      ReacTi : G7_TransitionPlus_V6;   // Transition structure
      ReacD : G7_TransitionPlus_V6;   // Transition structure
      Confirm : G7_TransitionPlus_V6;   // Transition structure
      UserBtch : G7_TransitionPlus_V6;   // Transition structure
      "StT-103" : G7_TransitionPlus_V6;   // Transition structure
      Route_Ok : G7_TransitionPlus_V6;   // Transition structure
      MixDone : G7_TransitionPlus_V6;   // Transition structure
      TimeOut : G7_TransitionPlus_V6;   // Transition structure
      EmptyLv : G7_TransitionPlus_V6;   // Transition structure
      LR : G7_TransitionPlus_V6;   // Transition structure
      LFUW : G7_TransitionPlus_V6;   // Transition structure
      mtL : G7_TransitionPlus_V6;   // Transition structure
      DneTransf : G7_TransitionPlus_V6;   // Transition structure
      TWash : G7_TransitionPlus_V6;   // Transition structure
      STW : G7_TransitionPlus_V6;   // Transition structure
      OpRout : G7_TransitionPlus_V6;   // Transition structure
      TW_RW : G7_TransitionPlus_V6;   // Transition structure
      TW_Vfd : G7_TransitionPlus_V6;   // Transition structure
      Trans87 : G7_TransitionPlus_V6;   // Transition structure
      TW_Wng : G7_TransitionPlus_V6;   // Transition structure
      TW_VfdOf : G7_TransitionPlus_V6;   // Transition structure
      Trans90 : G7_TransitionPlus_V6;   // Transition structure
      DneTnkW : G7_TransitionPlus_V6;   // Transition structure
      TE_SWW : G7_TransitionPlus_V6;   // Transition structure
      TuW : G7_TransitionPlus_V6;   // Transition structure
      STuW : G7_TransitionPlus_V6;   // Transition structure
      Trans103 : G7_TransitionPlus_V6;   // Transition structure
      TuWRW : G7_TransitionPlus_V6;   // Transition structure
      TuWGW : G7_TransitionPlus_V6;   // Transition structure
      TuW_SRW : G7_TransitionPlus_V6;   // Transition structure
      TuW_R : G7_TransitionPlus_V6;   // Transition structure
      Trans108 : G7_TransitionPlus_V6;   // Transition structure
      Trans109 : G7_TransitionPlus_V6;   // Transition structure
      PmpsOn : G7_TransitionPlus_V6;   // Transition structure
      ReEmpty : G7_TransitionPlus_V6;   // Transition structure
      PmpsOff : G7_TransitionPlus_V6;   // Transition structure
      OutleClsd : G7_TransitionPlus_V6;   // Transition structure
      DneTubW : G7_TransitionPlus_V6;   // Transition structure
      Init : G7_TransitionPlus_V6;   // Transition structure
      SAut : G7_TransitionPlus_V6;   // Transition structure
      SIn : G7_TransitionPlus_V6;   // Transition structure
      Initd : G7_TransitionPlus_V6;   // Transition structure
      WaterDn : G7_TransitionPlus_V6;   // Transition structure
      Ab : G7_TransitionPlus_V6;   // Transition structure
      AbortOn : G7_TransitionPlus_V6;   // Transition structure
      DneAbort : G7_TransitionPlus_V6;   // Transition structure
      Idle : G7_StepPlus_V6;   // Step structure
      Ready : G7_StepPlus_V6;   // Step structure
      SelectSeq : G7_StepPlus_V6;   // Step structure
      Started : G7_StepPlus_V6;   // Step structure
      StartTanks : G7_StepPlus_V6;   // Step structure
      FillingUpWater : G7_StepPlus_V6;   // Step structure
      StopReqWaterP : G7_StepPlus_V6;   // Step structure
      ReleaseWTank : G7_StepPlus_V6;   // Step structure
      "Pre-Mix" : G7_StepPlus_V6;   // Step structure
      OpenRoutes : G7_StepPlus_V6;   // Step structure
      X : G7_StepPlus_V6;   // Step structure
      FillDone_T101 : G7_StepPlus_V6;   // Step structure
      Close_T101 : G7_StepPlus_V6;   // Step structure
      "T-101_Done" : G7_StepPlus_V6;   // Step structure
      Y : G7_StepPlus_V6;   // Step structure
      pH_Ctrl1 : G7_StepPlus_V6;   // Step structure
      pH_Ctrl2 : G7_StepPlus_V6;   // Step structure
      FillDone_T102 : G7_StepPlus_V6;   // Step structure
      Close_T102 : G7_StepPlus_V6;   // Step structure
      "T-102_Done" : G7_StepPlus_V6;   // Step structure
      ReactingTime : G7_StepPlus_V6;   // Step structure
      ReactingDone : G7_StepPlus_V6;   // Step structure
      "USER Waiting" : G7_StepPlus_V6;   // Step structure
      "EDIT BatchP" : G7_StepPlus_V6;   // Step structure
      "Start T-103" : G7_StepPlus_V6;   // Step structure
      "R-201-->T-103" : G7_StepPlus_V6;   // Step structure
      MixToClean : G7_StepPlus_V6;   // Step structure
      LastFlushOut : G7_StepPlus_V6;   // Step structure
      Transfering : G7_StepPlus_V6;   // Step structure
      LastFIllUp : G7_StepPlus_V6;   // Step structure
      FirstFlushOut : G7_StepPlus_V6;   // Step structure
      LastFillUpW : G7_StepPlus_V6;   // Step structure
      LastTransfer : G7_StepPlus_V6;   // Step structure
      Done_Transfer : G7_StepPlus_V6;   // Step structure
      Idle_TWash : G7_StepPlus_V6;   // Step structure
      Start_TWash : G7_StepPlus_V6;   // Step structure
      OpenRoute : G7_StepPlus_V6;   // Step structure
      ReqWaterWash : G7_StepPlus_V6;   // Step structure
      "2011 VFD ON & PID AUTO/Wait for 80%_R-201" : G7_StepPlus_V6;   // Step structure
      StopWaterWash : G7_StepPlus_V6;   // Step structure
      "XV-1043_CC_02_R-201" : G7_StepPlus_V6;   // Step structure
      Washing : G7_StepPlus_V6;   // Step structure
      "2011VFD OFF & PID MAN_R-201" : G7_StepPlus_V6;   // Step structure
      USER_MAN_DRAIN : G7_StepPlus_V6;   // Step structure
      Done_TWash : G7_StepPlus_V6;   // Step structure
      Idle_TubWash : G7_StepPlus_V6;   // Step structure
      Start_TubWash : G7_StepPlus_V6;   // Step structure
      "XV-1043_CO_03_R-201" : G7_StepPlus_V6;   // Step structure
      ReqWaterTuW : G7_StepPlus_V6;   // Step structure
      GettingWater : G7_StepPlus_V6;   // Step structure
      StopRqWaterTuW : G7_StepPlus_V6;   // Step structure
      "ReleaseT-104" : G7_StepPlus_V6;   // Step structure
      "XV-1043_CC_03_R-529" : G7_StepPlus_V6;   // Step structure
      "XV-2013_CO_XV-1043_Cc_R-201" : G7_StepPlus_V6;   // Step structure
      "P-201A/B_ON_R-201" : G7_StepPlus_V6;   // Step structure
      Emptying : G7_StepPlus_V6;   // Step structure
      "P-201A/B_OFF_R-201" : G7_StepPlus_V6;   // Step structure
      Close_Outlet : G7_StepPlus_V6;   // Step structure
      Done_TubWash : G7_StepPlus_V6;   // Step structure
      Initialize : G7_StepPlus_V6;   // Step structure
      SetAuto : G7_StepPlus_V6;   // Step structure
      SetInitial : G7_StepPlus_V6;   // Step structure
      Initialized : G7_StepPlus_V6;   // Step structure
      AbortStarting : G7_StepPlus_V6;   // Step structure
      Aborting : G7_StepPlus_V6;   // Step structure
      Abort_Done : G7_StepPlus_V6;   // Step structure
      SINI : Array[0..9] of USInt;
      LSTT : Array[0..68] of USInt;
      ATAJ : Array[0..68] of USInt;
      ATAB : Array[0..68] of USInt;
      PSTT : Array[0..68] of USInt;
      NSTT : Array[0..68] of USInt;
      ASSJ : Array[0..65] of USInt;
      ASSB : Array[0..65] of USInt;
      PTTS : Array[0..65] of USInt;
      NTTS : Array[0..65] of USInt;
      SW_SQTS : Array[0..65] of USInt;
      SWITCH : Array[0..15] of USInt;
      TVX : Array[0..15] of USInt;
      TTX : Array[0..15] of USInt;
      TSX : Array[0..9] of USInt;
      S00X : Array[0..9] of USInt;
      SOFFX : Array[0..9] of USInt;
      SONX : Array[0..9] of USInt;
      SAX : Array[0..9] of USInt;
      SERRX : Array[0..66] of USInt;
      SMX : Array[0..66] of USInt;
      S0X : Array[0..66] of USInt;
      S1X : Array[0..66] of USInt;
      IL_ALARM_INST : Diag_Alarm;
      SUP_ALARM_INST : Diag_Alarm;
      STEP_TIME_ALARM_INST : Diag_Alarm;
      IEC_TIMER_INST : IEC_TIMER;
      TRANSACTION_FLAG : Bool := false;
   END_VAR
   VAR CONSTANT
      "Single R-201 T-101 seq done" : Int := 214;
      "Single R-201 T-102 seq done" : Int := 218;
   END_VAR
   // SINI[0] := 2;
   // LSTT[0] := 63;
   // NSTT[0] := 63;
   // PTTS[0] := 255;
   // TVX[0] := 16#1;
   // TTX[0] := 16#1;
   // TSX[0] := 16#1;
   // S00X[0] := 16#1;
   // SOFFX[0] := 16#1;
   // SONX[0] := 16#1;
   // SAX[0] := 16#1;
   // SERRX[0] := 16#1;
   // SMX[0] := 16#1;
   // S0X[0] := 16#1;
   // S1X[0] := 16#1;
   // LSTT[38] := 255;
   // SINI[3] := 255;
   // LSTT[1] := 59;
   // LSTT[2] := 255;
   // LSTT[3] := 255;
   // LSTT[4] := 3;
   // LSTT[5] := 34;
   // LSTT[6] := 45;
   // LSTT[7] := 255;
   // LSTT[8] := 255;
   // LSTT[9] := 255;
   // LSTT[10] := 255;
   // LSTT[11] := 255;
   // LSTT[12] := 255;
   // LSTT[13] := 255;
   // LSTT[14] := 255;
   // LSTT[15] := 255;
   // LSTT[16] := 255;
   // LSTT[17] := 255;
   // LSTT[18] := 255;
   // LSTT[19] := 255;
   // LSTT[20] := 255;
   // LSTT[21] := 255;
   // LSTT[22] := 255;
   // LSTT[23] := 255;
   // LSTT[24] := 255;
   // LSTT[56] := 255;
   // LSTT[27] := 255;
   // LSTT[57] := 255;
   // LSTT[29] := 255;
   // LSTT[30] := 255;
   // LSTT[31] := 255;
   // LSTT[32] := 255;
   // LSTT[55] := 255;
   // LSTT[62] := 255;
   // LSTT[44] := 255;
   // LSTT[36] := 255;
   // LSTT[66] := 255;
   // LSTT[39] := 255;
   // LSTT[40] := 255;
   // LSTT[41] := 255;
   // LSTT[42] := 255;
   // LSTT[59] := 255;
   // LSTT[58] := 255;
   // LSTT[46] := 255;
   // LSTT[47] := 255;
   // LSTT[50] := 255;
   // LSTT[51] := 255;
   // LSTT[52] := 255;
   // LSTT[53] := 255;
   // LSTT[54] := 255;
   // NSTT[28] := 28;
   // NSTT[65] := 33;
   // ATAJ[1] := 1;
   // ATAJ[2] := 2;
   // ATAJ[3] := 3;
   // ATAJ[4] := 4;
   // ATAJ[5] := 5;
   // ATAJ[6] := 6;
   // ATAJ[7] := 7;
   // ATAJ[8] := 8;
   // ATAJ[9] := 9;
   // ATAJ[10] := 10;
   // ATAJ[11] := 11;
   // ATAJ[12] := 12;
   // ATAJ[13] := 13;
   // ATAJ[14] := 14;
   // ATAJ[15] := 15;
   // ATAJ[16] := 16;
   // ATAJ[17] := 17;
   // ATAJ[18] := 18;
   // ATAJ[19] := 19;
   // ATAJ[20] := 20;
   // ATAJ[21] := 21;
   // ATAJ[22] := 22;
   // ATAJ[23] := 23;
   // ATAJ[24] := 24;
   // ATAJ[25] := 25;
   // ATAJ[26] := 26;
   // ATAJ[27] := 27;
   // ATAJ[28] := 28;
   // ATAJ[29] := 29;
   // ATAJ[30] := 30;
   // ATAJ[31] := 31;
   // ATAJ[32] := 32;
   // ATAJ[33] := 33;
   // ATAJ[34] := 34;
   // ATAJ[35] := 35;
   // ATAJ[36] := 36;
   // ATAJ[37] := 37;
   // ATAJ[38] := 38;
   // ATAJ[39] := 39;
   // ATAJ[40] := 40;
   // ATAJ[41] := 41;
   // ATAJ[42] := 42;
   // ATAJ[43] := 43;
   // ATAJ[44] := 44;
   // ATAJ[45] := 45;
   // ATAJ[46] := 46;
   // ATAJ[47] := 47;
   // ATAJ[48] := 48;
   // ATAJ[49] := 49;
   // ATAJ[50] := 50;
   // ATAJ[51] := 51;
   // ATAJ[52] := 52;
   // ATAJ[53] := 53;
   // ATAJ[54] := 54;
   // ATAJ[55] := 55;
   // ATAJ[56] := 56;
   // ATAJ[57] := 57;
   // ATAJ[58] := 58;
   // ATAJ[59] := 59;
   // ATAJ[60] := 60;
   // ATAJ[61] := 61;
   // ATAJ[62] := 62;
   // ATAJ[63] := 63;
   // ATAJ[64] := 64;
   // ATAJ[65] := 65;
   // ATAB[1] := 2;
   // ATAB[24] := 24;
   // ATAB[3] := 3;
   // ATAB[4] := 5;
   // ATAB[5] := 6;
   // ATAB[6] := 4;
   // ATAB[7] := 7;
   // ATAB[8] := 8;
   // ATAB[9] := 9;
   // ATAB[10] := 10;
   // ATAB[11] := 11;
   // ATAB[12] := 12;
   // ATAB[13] := 13;
   // ATAB[14] := 14;
   // ATAB[15] := 15;
   // ATAB[16] := 16;
   // ATAB[17] := 17;
   // ATAB[18] := 18;
   // ATAB[21] := 21;
   // ATAB[22] := 22;
   // ATAB[23] := 23;
   // ATAB[29] := 29;
   // ATAB[25] := 25;
   // ATAB[26] := 26;
   // ATAB[27] := 27;
   // ATAB[28] := 28;
   // ATAB[30] := 30;
   // ATAB[31] := 31;
   // ATAB[32] := 32;
   // ATAB[33] := 33;
   // ATAB[34] := 34;
   // ATAB[35] := 35;
   // ATAB[36] := 36;
   // ATAB[37] := 37;
   // ATAB[38] := 38;
   // ATAB[39] := 39;
   // ATAB[40] := 40;
   // ATAB[41] := 41;
   // ATAB[42] := 42;
   // ATAB[43] := 43;
   // ATAB[44] := 44;
   // ATAB[45] := 45;
   // ATAB[46] := 46;
   // ATAB[47] := 47;
   // ATAB[48] := 48;
   // ATAB[49] := 49;
   // ATAB[50] := 50;
   // ATAB[51] := 51;
   // ATAB[52] := 52;
   // ATAB[53] := 53;
   // ATAB[54] := 54;
   // ATAB[55] := 55;
   // ATAB[56] := 56;
   // ATAB[57] := 57;
   // ATAB[58] := 58;
   // ATAB[59] := 59;
   // ATAB[60] := 60;
   // ATAB[61] := 61;
   // ATAB[62] := 62;
   // ATAB[63] := 63;
   // ATAB[64] := 64;
   // ATAB[65] := 65;
   // PSTT[33] := 31;
   // PSTT[16] := 12;
   // PSTT[3] := 1;
   // PSTT[4] := 2;
   // PSTT[5] := 2;
   // PSTT[6] := 2;
   // PSTT[7] := 3;
   // PSTT[8] := 4;
   // PSTT[9] := 5;
   // PSTT[10] := 6;
   // PSTT[12] := 8;
   // PSTT[13] := 9;
   // PSTT[60] := 58;
   // PSTT[14] := 10;
   // PSTT[17] := 14;
   // PSTT[18] := 15;
   // PSTT[19] := 16;
   // PSTT[20] := 17;
   // PSTT[21] := 18;
   // PSTT[22] := 13;
   // PSTT[23] := 20;
   // PSTT[24] := 21;
   // PSTT[25] := 22;
   // PSTT[26] := 23;
   // PSTT[27] := 24;
   // PSTT[28] := 25;
   // PSTT[29] := 26;
   // PSTT[30] := 27;
   // PSTT[31] := 28;
   // PSTT[32] := 30;
   // PSTT[40] := 38;
   // PSTT[38] := 36;
   // PSTT[35] := 33;
   // PSTT[36] := 34;
   // PSTT[37] := 35;
   // PSTT[59] := 57;
   // PSTT[41] := 40;
   // PSTT[58] := 56;
   // PSTT[42] := 41;
   // PSTT[43] := 42;
   // PSTT[44] := 43;
   // PSTT[45] := 44;
   // PSTT[46] := 39;
   // PSTT[47] := 45;
   // PSTT[48] := 46;
   // PSTT[49] := 47;
   // PSTT[50] := 48;
   // PSTT[51] := 49;
   // PSTT[52] := 50;
   // PSTT[56] := 54;
   // PSTT[57] := 55;
   // PSTT[61] := 59;
   // PSTT[62] := 60;
   // PSTT[63] := 61;
   // PSTT[64] := 62;
   // PSTT[65] := 29;
   // NSTT[1] := 59;
   // NSTT[2] := 1;
   // NSTT[3] := 2;
   // NSTT[4] := 3;
   // NSTT[5] := 34;
   // NSTT[6] := 45;
   // NSTT[7] := 23;
   // NSTT[8] := 5;
   // NSTT[9] := 6;
   // NSTT[10] := 7;
   // NSTT[11] := 8;
   // NSTT[12] := 9;
   // NSTT[13] := 10;
   // NSTT[14] := 11;
   // NSTT[15] := 12;
   // NSTT[16] := 13;
   // NSTT[17] := 15;
   // NSTT[18] := 16;
   // NSTT[19] := 17;
   // NSTT[20] := 18;
   // NSTT[21] := 19;
   // NSTT[22] := 20;
   // NSTT[23] := 21;
   // NSTT[24] := 22;
   // NSTT[56] := 55;
   // NSTT[27] := 25;
   // NSTT[57] := 56;
   // NSTT[29] := 32;
   // NSTT[30] := 29;
   // NSTT[31] := 30;
   // NSTT[32] := 31;
   // NSTT[55] := 54;
   // NSTT[62] := 61;
   // NSTT[44] := 44;
   // NSTT[36] := 35;
   // NSTT[66] := 64;
   // NSTT[39] := 38;
   // NSTT[40] := 39;
   // NSTT[41] := 41;
   // NSTT[42] := 42;
   // NSTT[59] := 58;
   // NSTT[58] := 57;
   // NSTT[46] := 40;
   // NSTT[47] := 46;
   // NSTT[50] := 49;
   // NSTT[51] := 50;
   // NSTT[52] := 51;
   // NSTT[53] := 52;
   // NSTT[54] := 53;
   // LSTT[65] := 255;
   // ASSJ[1] := 1;
   // ASSJ[2] := 2;
   // ASSJ[3] := 3;
   // ASSJ[4] := 4;
   // ASSJ[5] := 5;
   // ASSJ[6] := 6;
   // ASSJ[7] := 7;
   // ASSJ[8] := 8;
   // ASSJ[9] := 9;
   // ASSJ[10] := 10;
   // ASSJ[11] := 11;
   // ASSJ[12] := 12;
   // ASSJ[13] := 19;
   // ASSJ[14] := 14;
   // ASSJ[15] := 15;
   // ASSJ[16] := 16;
   // ASSJ[17] := 17;
   // ASSJ[18] := 18;
   // ASSJ[19] := 13;
   // ASSJ[20] := 20;
   // ASSJ[21] := 21;
   // ASSJ[22] := 22;
   // ASSJ[23] := 23;
   // ASSJ[24] := 24;
   // ASSJ[25] := 25;
   // ASSJ[26] := 26;
   // ASSJ[27] := 27;
   // ASSJ[28] := 28;
   // ASSJ[29] := 29;
   // ASSJ[30] := 30;
   // ASSJ[31] := 31;
   // ASSJ[32] := 32;
   // ASSJ[33] := 33;
   // ASSJ[34] := 34;
   // ASSJ[35] := 35;
   // ASSJ[36] := 36;
   // ASSJ[37] := 37;
   // ASSJ[38] := 38;
   // ASSJ[39] := 39;
   // ASSJ[40] := 40;
   // ASSJ[41] := 41;
   // ASSJ[42] := 42;
   // ASSJ[43] := 43;
   // ASSJ[44] := 44;
   // ASSJ[45] := 45;
   // ASSJ[46] := 46;
   // ASSJ[47] := 47;
   // ASSJ[48] := 48;
   // ASSJ[49] := 49;
   // ASSJ[50] := 50;
   // ASSJ[51] := 51;
   // ASSJ[52] := 52;
   // ASSJ[53] := 53;
   // ASSJ[54] := 54;
   // ASSJ[55] := 55;
   // ASSJ[56] := 56;
   // ASSJ[57] := 57;
   // ASSJ[58] := 58;
   // ASSJ[59] := 59;
   // ASSJ[60] := 60;
   // ASSJ[61] := 61;
   // ASSJ[62] := 62;
   // ASSJ[63] := 63;
   // ASSB[1] := 1;
   // ASSB[2] := 2;
   // ASSB[3] := 3;
   // ASSB[4] := 4;
   // ASSB[5] := 5;
   // ASSB[6] := 6;
   // ASSB[7] := 7;
   // ASSB[8] := 8;
   // ASSB[9] := 9;
   // ASSB[10] := 14;
   // ASSB[11] := 11;
   // ASSB[12] := 12;
   // ASSB[13] := 13;
   // ASSB[14] := 10;
   // ASSB[15] := 15;
   // ASSB[16] := 16;
   // ASSB[17] := 17;
   // ASSB[18] := 18;
   // ASSB[19] := 19;
   // ASSB[20] := 20;
   // ASSB[21] := 21;
   // ASSB[22] := 22;
   // ASSB[23] := 23;
   // ASSB[24] := 24;
   // ASSB[25] := 25;
   // ASSB[26] := 26;
   // ASSB[27] := 27;
   // ASSB[28] := 28;
   // ASSB[29] := 29;
   // ASSB[30] := 30;
   // ASSB[31] := 31;
   // ASSB[32] := 32;
   // ASSB[33] := 33;
   // ASSB[34] := 34;
   // ASSB[35] := 35;
   // ASSB[36] := 36;
   // ASSB[37] := 37;
   // ASSB[38] := 38;
   // ASSB[39] := 39;
   // ASSB[40] := 40;
   // ASSB[41] := 41;
   // ASSB[42] := 42;
   // ASSB[43] := 43;
   // ASSB[44] := 44;
   // ASSB[45] := 45;
   // ASSB[46] := 46;
   // ASSB[47] := 47;
   // ASSB[48] := 48;
   // ASSB[49] := 49;
   // ASSB[50] := 50;
   // ASSB[51] := 51;
   // ASSB[52] := 52;
   // ASSB[53] := 53;
   // ASSB[54] := 54;
   // ASSB[55] := 55;
   // ASSB[56] := 56;
   // ASSB[57] := 57;
   // ASSB[58] := 58;
   // ASSB[59] := 59;
   // ASSB[60] := 60;
   // ASSB[61] := 61;
   // ASSB[62] := 62;
   // ASSB[63] := 63;
   // PTTS[3] := 255;
   // PTTS[61] := 62;
   // PTTS[5] := 8;
   // PTTS[6] := 9;
   // PTTS[7] := 10;
   // PTTS[8] := 11;
   // PTTS[9] := 12;
   // PTTS[10] := 13;
   // PTTS[11] := 14;
   // PTTS[12] := 15;
   // PTTS[13] := 16;
   // PTTS[14] := 13;
   // PTTS[15] := 17;
   // PTTS[16] := 18;
   // PTTS[17] := 19;
   // PTTS[18] := 20;
   // PTTS[19] := 21;
   // PTTS[20] := 22;
   // PTTS[21] := 23;
   // PTTS[22] := 24;
   // PTTS[23] := 7;
   // PTTS[24] := 255;
   // PTTS[25] := 27;
   // PTTS[26] := 33;
   // SW_SQTS[3] := 2;
   // PTTS[31] := 32;
   // PTTS[32] := 29;
   // PTTS[33] := 65;
   // PTTS[34] := 255;
   // PTTS[35] := 36;
   // PTTS[36] := 37;
   // PTTS[37] := 38;
   // PTTS[38] := 39;
   // PTTS[39] := 40;
   // PTTS[40] := 46;
   // PTTS[41] := 41;
   // PTTS[42] := 42;
   // PTTS[43] := 43;
   // PTTS[44] := 44;
   // PTTS[45] := 255;
   // PTTS[46] := 47;
   // PTTS[47] := 48;
   // PTTS[48] := 49;
   // PTTS[49] := 50;
   // PTTS[50] := 51;
   // PTTS[51] := 52;
   // PTTS[52] := 53;
   // PTTS[53] := 54;
   // PTTS[54] := 55;
   // PTTS[55] := 56;
   // PTTS[56] := 57;
   // PTTS[57] := 58;
   // PTTS[58] := 59;
   // PTTS[59] := 255;
   // PTTS[60] := 61;
   // SW_SQTS[34] := 7;
   // PTTS[62] := 63;
   // PTTS[63] := 255;
   // SW_SQTS[35] := 7;
   // NTTS[3] := 7;
   // NTTS[5] := 9;
   // NTTS[6] := 10;
   // NTTS[7] := 11;
   // NTTS[8] := 12;
   // NTTS[9] := 13;
   // NTTS[10] := 14;
   // NTTS[11] := 15;
   // NTTS[12] := 16;
   // NTTS[13] := 22;
   // NTTS[14] := 17;
   // NTTS[15] := 18;
   // NTTS[16] := 19;
   // NTTS[17] := 20;
   // NTTS[18] := 21;
   // NTTS[19] := 22;
   // NTTS[20] := 23;
   // NTTS[21] := 24;
   // NTTS[22] := 25;
   // NTTS[23] := 26;
   // NTTS[24] := 27;
   // NTTS[25] := 28;
   // NTTS[26] := 29;
   // NTTS[27] := 30;
   // NTTS[28] := 31;
   // NTTS[29] := 65;
   // NTTS[30] := 32;
   // NTTS[31] := 33;
   // NTTS[32] := 34;
   // NTTS[33] := 35;
   // NTTS[34] := 36;
   // NTTS[35] := 37;
   // NTTS[36] := 38;
   // NTTS[37] := 39;
   // NTTS[38] := 40;
   // NTTS[39] := 46;
   // NTTS[40] := 41;
   // NTTS[41] := 42;
   // NTTS[42] := 43;
   // NTTS[43] := 44;
   // NTTS[44] := 45;
   // NTTS[45] := 47;
   // NTTS[46] := 48;
   // NTTS[47] := 49;
   // NTTS[48] := 50;
   // NTTS[49] := 51;
   // NTTS[50] := 52;
   // NTTS[51] := 53;
   // NTTS[52] := 54;
   // NTTS[53] := 55;
   // NTTS[54] := 56;
   // NTTS[55] := 57;
   // NTTS[56] := 58;
   // NTTS[57] := 59;
   // NTTS[58] := 60;
   // NTTS[59] := 61;
   // NTTS[60] := 62;
   // NTTS[61] := 63;
   // NTTS[62] := 64;
   // NTTS[63] := 66;
   // SW_SQTS[2] := 1;
   // SW_SQTS[8] := 2;
   // SW_SQTS[9] := 2;
   // SW_SQTS[10] := 3;
   // SW_SQTS[11] := 3;
   // SW_SQTS[12] := 3;
   // SW_SQTS[13] := 3;
   // SW_SQTS[14] := 4;
   // SW_SQTS[15] := 4;
   // SW_SQTS[16] := 4;
   // SW_SQTS[17] := 4;
   // SW_SQTS[18] := 4;
   // SW_SQTS[19] := 4;
   // SW_SQTS[20] := 5;
   // SW_SQTS[21] := 5;
   // SW_SQTS[22] := 5;
   // SW_SQTS[23] := 2;
   // SW_SQTS[24] := 6;
   // SW_SQTS[25] := 6;
   // SW_SQTS[26] := 6;
   // SW_SQTS[27] := 6;
   // SW_SQTS[28] := 6;
   // SW_SQTS[29] := 6;
   // SW_SQTS[30] := 6;
   // SW_SQTS[31] := 6;
   // SWITCH[3] := 240;
   // SW_SQTS[36] := 7;
   // SW_SQTS[37] := 7;
   // SW_SQTS[38] := 7;
   // SW_SQTS[39] := 7;
   // SW_SQTS[40] := 7;
   // SW_SQTS[41] := 7;
   // SW_SQTS[42] := 7;
   // SW_SQTS[43] := 7;
   // SW_SQTS[44] := 7;
   // SW_SQTS[45] := 8;
   // SW_SQTS[46] := 8;
   // SW_SQTS[47] := 8;
   // SW_SQTS[48] := 8;
   // SW_SQTS[49] := 8;
   // SW_SQTS[50] := 8;
   // SW_SQTS[51] := 8;
   // SW_SQTS[52] := 8;
   // SW_SQTS[53] := 8;
   // SW_SQTS[54] := 8;
   // SW_SQTS[55] := 8;
   // SW_SQTS[56] := 8;
   // SW_SQTS[57] := 8;
   // SW_SQTS[58] := 8;
   // SW_SQTS[59] := 9;
   // SW_SQTS[60] := 9;
   // SW_SQTS[61] := 9;
   // SW_SQTS[62] := 9;
   // SW_SQTS[63] := 10;
   // SWITCH[0] := 252;
   // SWITCH[8] := 255;
   // SWITCH[4] := 167;
   // SWITCH[5] := 191;
   // SWITCH[6] := 252;
   // SWITCH[7] := 225;
   // SWITCH[2] := 255;
   // NSTT[48] := 47;
   // PTTS[27] := 34;
   // NSTT[38] := 37;
   // PTTS[30] := 31;
   // NTTS[1] := 3;
   // SWITCH[14] := 255;
   // ATAB[67] := 67;
   // ATAB[20] := 20;
   // PSTT[11] := 7;
   // NTTS[2] := 4;
   // PTTS[4] := 26;
   // PTTS[1] := 2;
   // PSTT[67] := 64;
   // NTTS[4] := 8;
   // ATAJ[67] := 67;
   // SW_SQTS[1] := 1;
   // NSTT[26] := 4;
   // LSTT[48] := 255;
   // LSTT[63] := 255;
   // NSTT[63] := 62;
   // LSTT[61] := 255;
   // NSTT[61] := 60;
   // LSTT[64] := 1;
   // NSTT[64] := 1;
   // "Aux Reactor"."TIMER".MIX.PT := T#5M;
   // "Aux Reactor"."TIMER"."PRE-MIX".PT := T#5M;
   // SINI[6] := 255;
   // "Aux Reactor"."TIMER".TUBE.PT := T#5M;
   // "Aux Reactor"."TIMER".WASH.PT := T#5M;
   // SINI[5] := 255;
   // "Aux Reactor"."TIMER".REACTOR.PT := T#21.5H;
   // "Aux Reactor"."TIMER".PH_DELAY.PT := T#1M;
   // PTTS[29] := 30;
   // LSTT[37] := 255;
   // LSTT[25] := 24;
   // ATAB[19] := 19;
   // PSTT[15] := 11;
   // NSTT[37] := 36;
   // NSTT[25] := 24;
   // PTTS[28] := 28;
   // SW_SQTS[7] := 2;
   // SW_SQTS[6] := 2;
   // SW_SQTS[5] := 2;
   // SW_SQTS[4] := 2;
   // SWITCH[11] := 255;
   // SWITCH[13] := 239;
   // SWITCH[12] := 254;
   // PSTT[34] := 32;
   // PSTT[55] := 53;
   // PSTT[54] := 52;
   // LSTT[26] := 255;
   // SWITCH[10] := 239;
   // SWITCH[9] := 254;
   // SWITCH[1] := 231;
   // PTTS[2] := 3;
   // NSTT[49] := 48;
   // PSTT[53] := 51;
   // ATAB[0] := 1;
   // LSTT[49] := 255;
   // SINI[4] := 255;
   // SINI[2] := 255;
   // SW_SQTS[33] := 6;
   // SW_SQTS[32] := 6;
   // NSTT[34] := 27;
   // SINI[7] := 255;
   // SINI[8] := 255;
   // SINI[9] := 255;
   // LSTT[34] := 255;
   // LSTT[43] := 255;
   // PSTT[39] := 37;
   // NSTT[43] := 43;
   // LSTT[28] := 255;
   // LSTT[33] := 255;
   // ATAJ[66] := 66;
   // ATAB[66] := 66;
   // PSTT[66] := 63;
   // NSTT[33] := 26;
   // ASSJ[64] := 64;
   // ASSB[64] := 64;
   // PTTS[64] := 66;
   // NTTS[64] := 67;
   // SW_SQTS[64] := 10;
   // LSTT[67] := 255;
   // ATAJ[68] := 68;
   // ATAB[68] := 68;
   // PSTT[68] := 65;
   // NSTT[67] := 65;
   // ASSJ[65] := 65;
   // ASSB[65] := 65;
   // PTTS[65] := 67;
   // NTTS[65] := 68;
   // SW_SQTS[65] := 10;
BEGIN
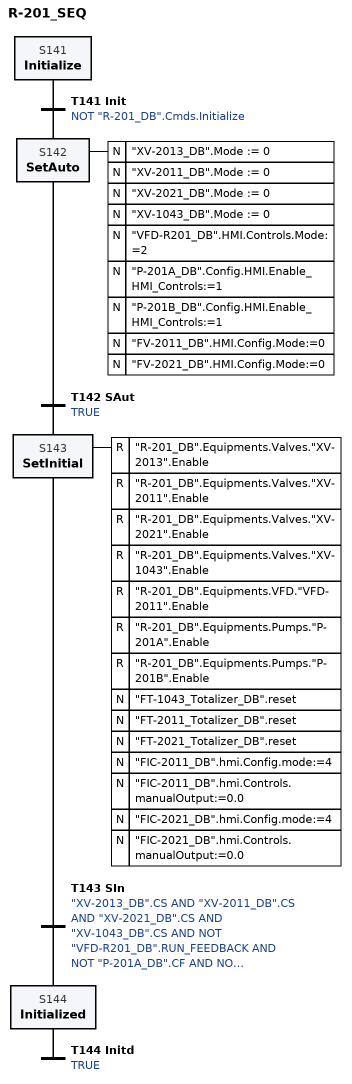
   // permanent pre-instructions
   NETWORK 1
      "R-201_Signals_FROM_T-101"();
      "R-201_Signals_FROM_T-102"();
      "R-201_Signals_FROM_T-103"();
      "R-201_Signals_FROM_T-104"();
      "R-201_SEQ_FC"();
      "R-201_Transitions_FC"();

   // sequencer 1
   STEP Initialize:   // S141, max time T#10S, warning time T#7S
   END_STEP
   TRANSITION Init FROM Initialize TO SetAuto   // T141
      := NOT "R-201_DB".Cmds.Initialize;
   END_TRANSITION
   STEP SetAuto:   // S142, max time T#10S, warning time T#7S
              N    "XV-2013_DB".Mode := 0
              N    "XV-2011_DB".Mode := 0
              N    "XV-2021_DB".Mode := 0
              N    "XV-1043_DB".Mode := 0
              N    "VFD-R201_DB".HMI.Controls.Mode:=2
              N    "P-201A_DB".Config.HMI.Enable_HMI_Controls:=1
              N    "P-201B_DB".Config.HMI.Enable_HMI_Controls:=1
              N    "FV-2011_DB".HMI.Config.Mode:=0
              N    "FV-2021_DB".HMI.Config.Mode:=0
   END_STEP
   TRANSITION SAut FROM SetAuto TO SetInitial   // T142
      := TRUE;
   END_TRANSITION
   STEP SetInitial:   // S143, max time T#10S, warning time T#7S
              R    "R-201_DB".Equipments.Valves."XV-2013".Enable
              R    "R-201_DB".Equipments.Valves."XV-2011".Enable
              R    "R-201_DB".Equipments.Valves."XV-2021".Enable
              R    "R-201_DB".Equipments.Valves."XV-1043".Enable
              R    "R-201_DB".Equipments.VFD."VFD-2011".Enable
              R    "R-201_DB".Equipments.Pumps."P-201A".Enable
              R    "R-201_DB".Equipments.Pumps."P-201B".Enable
              N    "FT-1043_Totalizer_DB".reset
              N    "FT-2011_Totalizer_DB".reset
              N    "FT-2021_Totalizer_DB".reset
              N    "FIC-2011_DB".hmi.Config.mode:=4
              N    "FIC-2011_DB".hmi.Controls.manualOutput:=0.0
              N    "FIC-2021_DB".hmi.Config.mode:=4
              N    "FIC-2021_DB".hmi.Controls.manualOutput:=0.0
   END_STEP
   TRANSITION SIn FROM SetInitial TO Initialized   // T143
      := "XV-2013_DB".CS AND "XV-2011_DB".CS AND "XV-2021_DB".CS AND "XV-1043_DB".CS AND NOT "VFD-R201_DB".RUN_FEEDBACK AND NOT "P-201A_DB".CF AND NOT "P-201B_DB".CF AND ("FV-2011_DB".CMD <= 0) AND ("FV-2021_DB".CMD <= 0) AND ("FT-1043_Totalizer_DB".Total = 0.0) AND ("FT-2011_Totalizer_DB".Total = 0.0) AND ("FT-2021_Totalizer_DB".Total = 0.0);
   END_TRANSITION
   STEP Initialized:   // S144, max time T#10S, warning time T#7S
      // Done Initialization
   END_STEP
   TRANSITION Initd FROM Initialized TO ?   // T144
      := TRUE;
   END_TRANSITION

   // permanent post-instructions
   NETWORK 1
      "R-201_FC_Outputs"();
END_FUNCTION_BLOCK

FUNCTION "R-201_FC_Outputs" : Void   // FC36, SCL
{ S7_Optimized_Access := 'TRUE' }
VERSION : 0.1
   VAR_TEMP
      Pump_A : Struct
         Cond_01 : Bool;   // Condition 01
         Cond_02 : Bool;
         Cond_03 : Bool;   // Condition 03
      END_STRUCT;
      Pump_B : Struct
         Cond_01 : Bool;   // Condition 01
         Cond_02 : Bool;   // Condition 02
         Cond_03 : Bool;   // Condition 03
      END_STRUCT;
      Motor : Struct
         Cond_01 : Bool;   // Condition 01
         Cond_02 : Bool;   // Condition 02
         Cond_03 : Bool;   // Condition 03
      END_STRUCT;
      XV : Struct
         "2013" : Bool;
         "2011" : Bool;
         "2021" : Bool;
         "1043" : Bool;
      END_STRUCT;
      "FV-2011" : Struct
         On : Bool;
         Cond_1 : Bool;
      END_STRUCT;
      "FV-2021" : Struct
         On : Bool;
         Cond_1 : Bool;
      END_STRUCT;
   END_VAR
BEGIN
   //****** Equipmens Activation*******
   //
   //**************************************************************
   //
   //IF "AlwaysFALSE" THEN
       //***********************************************Reactor Outlet Valve**********************************************************************
       IF "XV-2013_DB".Mode = 0 THEN
           "R-201_DB".Equipments.Valves."XV-2013".CmdOn := "R-201_DB".Equipments.Valves."XV-2013".Enable AND NOT "R-201_DB".Cmds.Hold AND NOT "R-201_DB".Status.Aborting;
           //Delay Off To avoid Overpressure the Lines
           #XV."2013" := "R-201_DB".Equipments.Valves."XV-2013".CmdOn;
           "R-201_Aux_DB".Timer."XV-2013".TOF(IN := #XV."2013",
                                              PT := "R-201_Aux_DB".Constants.CmdDelay);
           //Command to the Valve
           IF "R-201_Aux_DB".Timer."XV-2013".Q THEN
               "XV-2013_DB".CMD := 2;
           ELSE
               "XV-2013_DB".CMD := 1;
           END_IF;
           "R-201_DB".Equipments.Valves."XV-2013".TurningOff := NOT "R-201_DB".Equipments.Valves."XV-2013".CmdOn AND "R-201_Aux_DB".Timer."XV-2013".Q;
       END_IF;
       //***********************************************From T-101 Inlet Route********************************************************************
       IF "XV-2011_DB".Mode = 0 THEN
           "R-201_DB".Equipments.Valves."XV-2011".CmdOn := "R-201_DB".Equipments.Valves."XV-2011".Enable AND NOT "R-201_DB".Cmds.Hold AND NOT "R-201_DB".Status.Aborting;
           //Delay Off To avoid Overpressure the Lines
           #XV."2011" := "R-201_DB".Equipments.Valves."XV-2011".CmdOn;
           "R-201_Aux_DB".Timer."XV-2011".TOF(IN := #XV."2011",
                                              PT := "R-201_Aux_DB".Constants.CmdDelay);
           //Command to the Valve
           IF "R-201_Aux_DB".Timer."XV-2011".Q THEN
               "XV-2011_DB".CMD := 2;
           ELSE
               "XV-2011_DB".CMD := 1;
           END_IF;
           "R-201_DB".Equipments.Valves."XV-2011".TurningOff := NOT "R-201_DB".Equipments.Valves."XV-2011".CmdOn AND "R-201_Aux_DB".Timer."XV-2011".Q;
       END_IF;
       //***********************************************From T-102 Inlet Route********************************************************************
       IF "XV-2021_DB".Mode = 0 THEN
           "R-201_DB".Equipments.Valves."XV-2021".CmdOn := "R-201_DB".Equipments.Valves."XV-2021".Enable AND NOT "R-201_DB".Cmds.Hold AND NOT "R-201_DB".Status.Aborting;
           //Delay Off To avoid Overpressure the Lines
           #XV."2021" := "R-201_DB".Equipments.Valves."XV-2021".CmdOn;
           "R-201_Aux_DB".Timer."XV-2021".TOF(IN := #XV."2021",
                                              PT := "R-201_Aux_DB".Constants.CmdDelay);
           IF "R-201_Aux_DB".Timer."XV-2021".Q THEN
               "XV-2021_DB".CMD := 2;
           ELSE
               "XV-2021_DB".CMD := 1;
           END_IF;
           "R-201_DB".Equipments.Valves."XV-2021".TurningOff := NOT "R-201_DB".Equipments.Valves."XV-2021".CmdOn AND "R-201_Aux_DB".Timer."XV-2021".Q;
       END_IF;
       //***********************************************From T-104 Inlet Route (Water)********************************************************************
       IF "XV-1043_DB".Mode = 0 THEN
           "R-201_DB".Equipments.Valves."XV-1043".CmdOn := "R-201_DB".Equipments.Valves."XV-1043".Enable AND NOT "R-201_DB".Cmds.Hold AND NOT "R-201_DB".Status.Aborting;
           //Delay Off To avoid Overpressure the Lines
           #XV."1043" := "R-201_DB".Equipments.Valves."XV-1043".CmdOn;
           "R-201_Aux_DB".Timer."XV-1043".TOF(IN := #XV."1043",
                                              PT := "R-201_Aux_DB".Constants.CmdDelay);
           IF "R-201_Aux_DB".Timer."XV-1043".Q THEN
               "XV-1043_DB".CMD := 2;
           ELSE
               "XV-1043_DB".CMD := 1;
           END_IF;
           "R-201_DB".Equipments.Valves."XV-1043".TurningOff := NOT "R-201_DB".Equipments.Valves."XV-1043".CmdOn AND "R-201_Aux_DB".Timer."XV-1043".Q;
       END_IF;
       //***********************************************FIC-2011 Controller (From T-101)********************************************************************
       IF "FV-2011_DB".HMI.Config.Mode=0 THEN
           #"FV-2011".Cond_1 := "R-201_DB".Equipments.Valves."FV-2011".Enable AND "XV-2011_DB".OS;
           "R-201_DB".Equipments.Valves."FV-2011".CmdOn := #"FV-2011".Cond_1 AND NOT "R-201_DB".Cmds.Hold AND NOT "R-201_DB".Status.Aborting;
           //Delay Off To avoid Overpressure the Lines
           #"FV-2011".On := "R-201_DB".Equipments.Valves."FV-2011".CmdOn;
           "R-201_Aux_DB".Timer."FV-2011".TOF(IN := #"FV-2011".On,
                                              PT := "R-201_Aux_DB".Constants.CmdDelay);
           IF "R-201_Aux_DB".Timer."FV-2011".Q THEN
               "FIC-2011_DB".enableManualMode := False;
               "FIC-2011_DB".enableRemoteSetpoint := False;
               "FIC-2011_DB".hmi.Controls.manualEnable := False;
               "FIC-2011_DB".hmi.Config.mode := 3;
           END_IF; //  ELSE
             //  "FIC-2011_DB".enableManualMode := True;
             //  "FIC-2011_DB".hmi.Controls.manualEnable := True;
            //   "FIC-2011_DB".hmi.Config.mode := 4;
             //  "FIC-2011_DB".hmi.Controls.manualOutput:=0;
          // END_IF;
           "R-201_DB".Equipments.Valves."FV-2011".TurningOff := NOT "R-201_DB".Equipments.Valves."FV-2011".CmdOn AND "R-201_Aux_DB".Timer."FV-2011".Q;
       END_IF;
       //***********************************************FIC-2021 Controller (From T-102)********************************************************************
       IF "FV-2021_DB".HMI.Config.Mode = 0 THEN
           #"FV-2021".Cond_1 := "R-201_DB".Equipments.Valves."FV-2021".Enable AND "XV-2021_DB".OS;
           "R-201_DB".Equipments.Valves."FV-2021".CmdOn := #"FV-2021".Cond_1 AND NOT "R-201_DB".Cmds.Hold AND NOT "R-201_DB".Status.Aborting;
           //Delay Off To avoid Overpressure the Lines
           #"FV-2021".On := "R-201_DB".Equipments.Valves."FV-2021".CmdOn;
           "R-201_Aux_DB".Timer."FV-2021".TOF(IN := #"FV-2021".On,
                                              PT := "R-201_Aux_DB".Constants.CmdDelay);
           IF "R-201_Aux_DB".Timer."FV-2021".Q THEN

               IF "R-201_SEQ_DB".pH_Ctrl1.X OR "R-201_SEQ_DB".pH_Ctrl2.X OR "R-201_SEQ_DB".FillDone_T102.X THEN
                   //FIC-2021 Secondary Controller
                   "FIC-2021_DB".enableManualMode := False;
                   "FIC-2021_DB".hmi.Controls.manualEnable := False;
                   "FIC-2021_DB".enableRemoteSetpoint := true;
                   "FIC-2021_DB".hmi.Config.mode := 6;

                   //PHIC-R-201 pH Primary Controller
                   "PHIC-R-201_DB".enableRemoteSetpoint := False;
                   "PHIC-R-201_DB".enableManualMode := False;
                   "PHIC-R-201_DB".hmi.Controls.manualEnable := False;
                   "PHIC-R-201_DB".hmi.Config.mode := 3;
               ELSIF "R-201_SEQ_DB".Y.X THEN
                   //FIC-2021 Secondary Controller
                   "FIC-2021_DB".enableManualMode := False;
                   "FIC-2021_DB".hmi.Controls.manualEnable := False;
                   "FIC-2021_DB".enableRemoteSetpoint := False;
                   "FIC-2021_DB".hmi.Config.mode := 3;

                   //PHIC-R-201 pH Primary Controller
                   "PHIC-R-201_DB".enableRemoteSetpoint := False;
                   "PHIC-R-201_DB".enableManualMode := False;
                   "PHIC-R-201_DB".hmi.Controls.manualEnable := False;
                   "PHIC-R-201_DB".hmi.Config.mode := 3;
               END_IF;

           END_IF; // ELSE
               //FIC-2021 Secondary Controller
              // "FIC-2011_DB".enableManualMode := True;
              // "FIC-2021_DB".hmi.Controls.manualEnable := True;
              // "FIC-2021_DB".enableRemoteSetpoint := False;
              // "FIC-2021_DB".hmi.Config.mode := 4;
              // "FIC-2021_DB".hmi.Controls.manualOutput := 0;

               //PHIC-R-201 pH Primary  Controller
              // "PHIC-R-201_DB".enableManualMode := True;
              // "PHIC-R-201_DB".hmi.Controls.manualEnable := True;
              // "PHIC-R-201_DB".enableRemoteSetpoint := False;
              // "PHIC-R-201_DB".hmi.Config.mode := 4;
              // "PHIC-R-201_DB".hmi.Controls.manualOutput := 0;


         //  END_IF;
           "R-201_DB".Equipments.Valves."FV-2021".TurningOff := NOT "R-201_DB".Equipments.Valves."FV-2021".CmdOn AND "R-201_Aux_DB".Timer."FV-2021".Q;
       END_IF;

       //***********************************************Recirculate/Feed Pump A********************************************************************
       // Condition to CmdOn "On Command" 
       IF "P-201A_DB".Config.HMI.Enable_HMI_Controls = 1 THEN
           #Pump_A.Cond_01 := "R-201_DB".Equipments.Pumps."P-201A".Enable AND ("R-201_DB".PmpSel."P-201AB" = 1 OR "R-201_DB".PmpSel."P-201AB" = 3);
           #Pump_A.Cond_02 := "XV-2013_DB".OS AND "R-201_Read_FROM_T-103_DB".RouteOpened; //Route Open to sent to the T-103 (Cooling Tank)
           "R-201_DB".Equipments.Pumps."P-201A".CmdOn := #Pump_A.Cond_01 AND #Pump_A.Cond_02 AND NOT "R-201_DB".Cmds.Hold AND NOT "R-201_DB".Status.Aborting;
           IF "R-201_DB".Equipments.Pumps."P-201A".CmdOn THEN
               "P-201A_DB".Stop_CMD := False;
               "P-201A_DB".Start_CMD := true;
               "P-201A_DB".ON := TRUE;
               "P-201A_DB".OFF := FALSE;
           ELSE
               "P-201A_DB".Stop_CMD := TRUE;
               "P-201A_DB".Start_CMD := FALSE;
               "P-201A_DB".ON := FALSE;
               "P-201A_DB".OFF := TRUE;
           END_IF;
       END_IF;
       //***********************************************Recirculate/Feed Pump B********************************************************************
       // Condition to CmdOn "On Command" 
       IF "P-201B_DB".Config.HMI.Enable_HMI_Controls = 1 THEN
           #Pump_B.Cond_01 := "R-201_DB".Equipments.Pumps."P-201B".Enable AND ("R-201_DB".PmpSel."P-201AB" = 2 OR "R-201_DB".PmpSel."P-201AB" = 3);
           #Pump_B.Cond_02 := "XV-2013_DB".OS AND "R-201_Read_FROM_T-103_DB".RouteOpened; //Route Open to sent to the T-103 (Cooling Tank)
           "R-201_DB".Equipments.Pumps."P-201B".CmdOn := #Pump_B.Cond_01 AND #Pump_B.Cond_02 AND NOT "R-201_DB".Cmds.Hold AND NOT "R-201_DB".Status.Aborting;
           IF "R-201_DB".Equipments.Pumps."P-201B".CmdOn THEN
               "P-201B_DB".Stop_CMD := False;
               "P-201B_DB".Start_CMD := true;
               "P-201B_DB".ON := TRUE;
               "P-201B_DB".OFF := FALSE;
           ELSE
               "P-201B_DB".Stop_CMD := TRUE;
               "P-201B_DB".Start_CMD := FALSE;
               "P-201B_DB".ON := FALSE;
               "P-201B_DB".OFF := TRUE;
           END_IF;
       END_IF;
       //***********************************************Mixer********************************************************************
       IF "VFD-R201_DB".HMI.Controls.Mode = 2 THEN
           "R-201_Aux_DB"."Real"."VFD-R201".Start := (("LT-2011_DB".SAI > "R-201_Recipe".MinLevelMixerOn+2.0)OR  "R-201_Aux_DB"."Real"."VFD-R201".Start) AND NOT "R-201_Aux_DB"."Real"."VFD-R201".Stop;
           "R-201_Aux_DB"."Real"."VFD-R201".Stop := ("LT-2011_DB".SAI < "R-201_Recipe".MinLevelMixerOn - 1.0);
           #Motor.Cond_01 := "R-201_DB".Equipments.VFD."VFD-2011".Enable AND  "R-201_Aux_DB"."Real"."VFD-R201".Start;
           "R-201_DB".Equipments.VFD."VFD-2011".CmdOn := #Motor.Cond_01 AND NOT "R-201_DB".Cmds.Hold AND NOT "R-201_DB".Status.Aborting;
           IF "R-201_DB".Equipments.VFD."VFD-2011".CmdOn THEN
               "VFD-R201_DB".PLCCommand := TRUE;
           ELSE
               "VFD-R201_DB".PLCCommand := FALSE;
           END_IF;
       END_IF;
   //END_IF;

   //***************Interlocks to T-103***************//
   //Transfering
   "R-201_Write_TO_T-103_DB".Transfering := ("XV-2013_DB".OS) AND (("P-201A_DB".CF AND ("PT-201A_DB".SAI > 0.2)) OR ("P-201B_DB".CF AND ("PT-201B_DB".SAI > 0.2)));
   "R-201_Write_TO_T-103_DB"."Transfer_To_T-103_Done" := "R-201_DB".Status.Step = 66;// AND "XV-2013_DB".CS AND NOT "P-201A_DB".CF AND NOT "P-201B_DB".CF AND NOT "VFD-R201_DB".RUN_FEEDBACK;
   //***************Interlocks to T-101***************//
   "R-201_Write_TO_T-101_DB".OpenRoute := "XV-2011_DB".OS AND ("FV-2011_DB".CMD > 0);
   "R-201_Write_TO_T-101_DB".RouteOpened := "XV-2011_DB".OS AND ("FV-2011_DB".CMD > 0);

   //***************Interlocks to T-102***************//
   "R-201_Write_TO_T-102_DB".OpenRoute := "XV-2021_DB".OS AND ("FV-2021_DB".CMD > 0);
   "R-201_Write_TO_T-102_DB".RouteOpened := "XV-2021_DB".OS AND ("FV-2021_DB".CMD > 0);
   //***************Abort Signals***************//
   //******Abort T-101*****//
   IF "R-201_DB".Status.Aborting THEN

